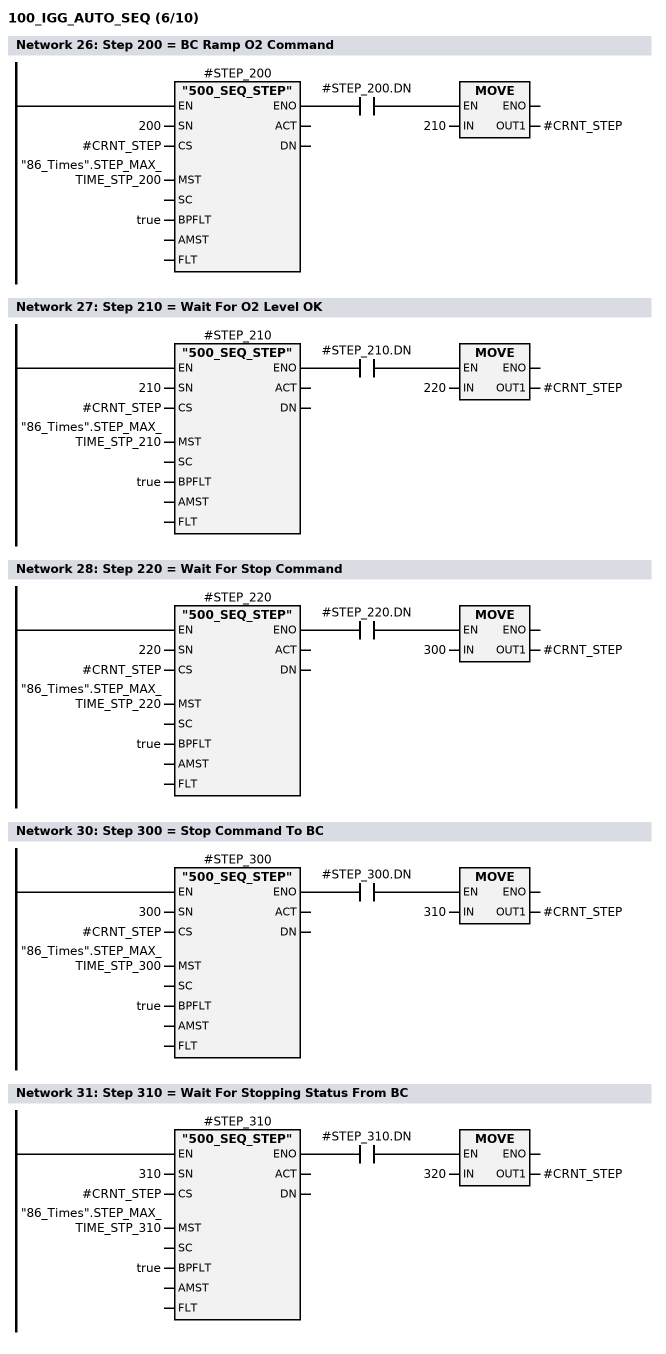
   RUNG wire#powerrail
      #STEP_200(SN := 200, CS := #CRNT_STEP, MST := "86_Times".STEP_MAX_TIME_STP_200, SC :=, BPFLT := true, AMST :=, FLT :=, ACT =>, DN =>)
      Contact( #STEP_200.DN )
      Move(in := 210, out1 => #CRNT_STEP)
   END_RUNG
   // the same network as SCL:
   #STEP_200(SN := 200, CS := #CRNT_STEP, MST := "86_Times".STEP_MAX_TIME_STP_200, BPFLT := true, ENO => #_w1);   // "500_SEQ_STEP"
   IF #_w1 AND #STEP_200.DN THEN #CRNT_STEP := 210; END_IF;
END_REGION

REGION Network 27: Step 210 = Wait For O2 Level OK
   RUNG wire#powerrail
      #STEP_210(SN := 210, CS := #CRNT_STEP, MST := "86_Times".STEP_MAX_TIME_STP_210, SC :=, BPFLT := true, AMST :=, FLT :=, ACT =>, DN =>)
      Contact( #STEP_210.DN )
      Move(in := 220, out1 => #CRNT_STEP)
   END_RUNG
   // the same network as SCL:
   #STEP_210(SN := 210, CS := #CRNT_STEP, MST := "86_Times".STEP_MAX_TIME_STP_210, BPFLT := true, ENO => #_w1);   // "500_SEQ_STEP"
   IF #_w1 AND #STEP_210.DN THEN #CRNT_STEP := 220; END_IF;
END_REGION

REGION Network 28: Step 220 = Wait For Stop Command
   RUNG wire#powerrail
      #STEP_220(SN := 220, CS := #CRNT_STEP, MST := "86_Times".STEP_MAX_TIME_STP_220, SC :=, BPFLT := true, AMST :=, FLT :=, ACT =>, DN =>)
      Contact( #STEP_220.DN )
      Move(in := 300, out1 => #CRNT_STEP)
   END_RUNG
   // the same network as SCL:
   #STEP_220(SN := 220, CS := #CRNT_STEP, MST := "86_Times".STEP_MAX_TIME_STP_220, BPFLT := true, ENO => #_w1);   // "500_SEQ_STEP"
   IF #_w1 AND #STEP_220.DN THEN #CRNT_STEP := 300; END_IF;
END_REGION

REGION Network 30: Step 300 = Stop Command To BC
   RUNG wire#powerrail
      #STEP_300(SN := 300, CS := #CRNT_STEP, MST := "86_Times".STEP_MAX_TIME_STP_300, SC :=, BPFLT := true, AMST :=, FLT :=, ACT =>, DN =>)
      Contact( #STEP_300.DN )
      Move(in := 310, out1 => #CRNT_STEP)
   END_RUNG
   // the same network as SCL:
   #STEP_300(SN := 300, CS := #CRNT_STEP, MST := "86_Times".STEP_MAX_TIME_STP_300, BPFLT := true, ENO => #_w1);   // "500_SEQ_STEP"
   IF #_w1 AND #STEP_300.DN THEN #CRNT_STEP := 310; END_IF;
END_REGION

REGION Network 31: Step 310 = Wait For Stopping Status From BC
   RUNG wire#powerrail
      #STEP_310(SN := 310, CS := #CRNT_STEP, MST := "86_Times".STEP_MAX_TIME_STP_310, SC :=, BPFLT := true, AMST :=, FLT :=, ACT =>, DN =>)
      Contact( #STEP_310.DN )
      Move(in := 320, out1 => #CRNT_STEP)
   END_RUNG
   // the same network as SCL:
   #STEP_310(SN := 310, CS := #CRNT_STEP, MST := "86_Times".STEP_MAX_TIME_STP_310, BPFLT := true, ENO => #_w1);   // "500_SEQ_STEP"
   IF #_w1 AND #STEP_310.DN THEN #CRNT_STEP := 320; END_IF;
END_REGION

REGION Network 32: Step 320 = Wait For O2 Control Stopped From BC
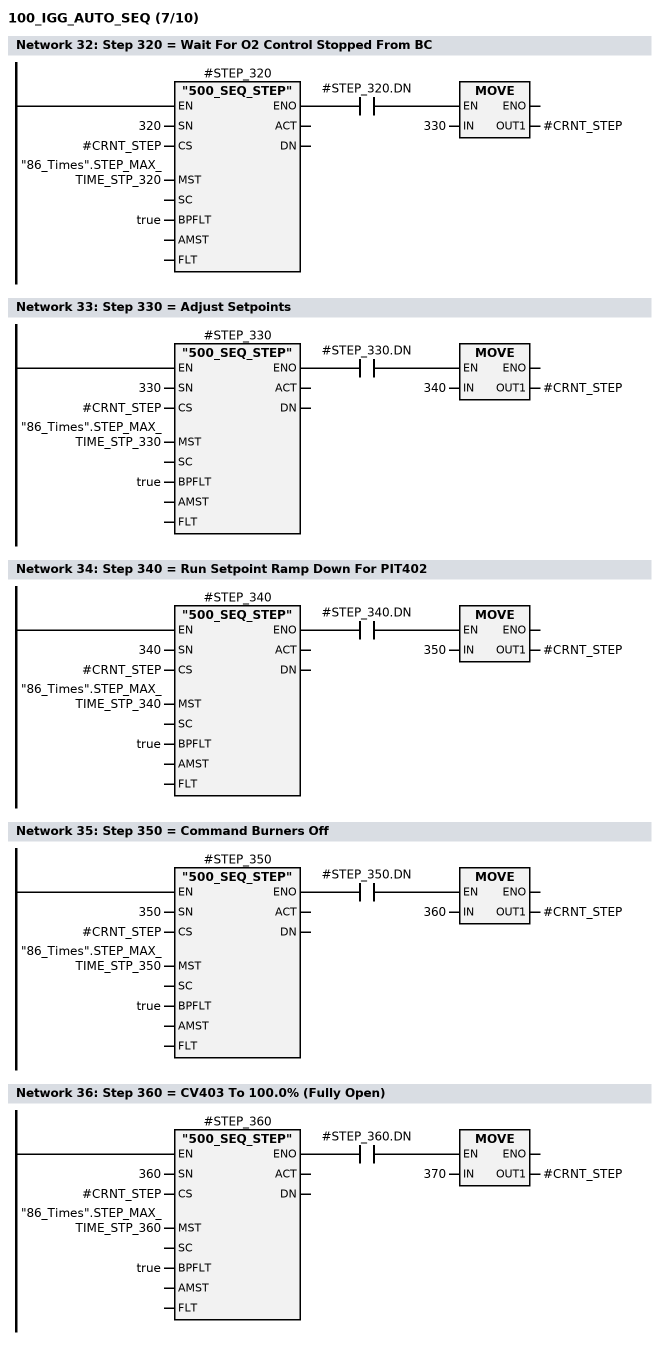
   RUNG wire#powerrail
      #STEP_320(SN := 320, CS := #CRNT_STEP, MST := "86_Times".STEP_MAX_TIME_STP_320, SC :=, BPFLT := true, AMST :=, FLT :=, ACT =>, DN =>)
      Contact( #STEP_320.DN )
      Move(in := 330, out1 => #CRNT_STEP)
   END_RUNG
   // the same network as SCL:
   #STEP_320(SN := 320, CS := #CRNT_STEP, MST := "86_Times".STEP_MAX_TIME_STP_320, BPFLT := true, ENO => #_w1);   // "500_SEQ_STEP"
   IF #_w1 AND #STEP_320.DN THEN #CRNT_STEP := 330; END_IF;
END_REGION

REGION Network 33: Step 330 = Adjust Setpoints
   RUNG wire#powerrail
      #STEP_330(SN := 330, CS := #CRNT_STEP, MST := "86_Times".STEP_MAX_TIME_STP_330, SC :=, BPFLT := true, AMST :=, FLT :=, ACT =>, DN =>)
      Contact( #STEP_330.DN )
      Move(in := 340, out1 => #CRNT_STEP)
   END_RUNG
   // the same network as SCL:
   #STEP_330(SN := 330, CS := #CRNT_STEP, MST := "86_Times".STEP_MAX_TIME_STP_330, BPFLT := true, ENO => #_w1);   // "500_SEQ_STEP"
   IF #_w1 AND #STEP_330.DN THEN #CRNT_STEP := 340; END_IF;
END_REGION

REGION Network 34: Step 340 = Run Setpoint Ramp Down For PIT402
   RUNG wire#powerrail
      #STEP_340(SN := 340, CS := #CRNT_STEP, MST := "86_Times".STEP_MAX_TIME_STP_340, SC :=, BPFLT := true, AMST :=, FLT :=, ACT =>, DN =>)
      Contact( #STEP_340.DN )
      Move(in := 350, out1 => #CRNT_STEP)
   END_RUNG
   // the same network as SCL:
   #STEP_340(SN := 340, CS := #CRNT_STEP, MST := "86_Times".STEP_MAX_TIME_STP_340, BPFLT := true, ENO => #_w1);   // "500_SEQ_STEP"
   IF #_w1 AND #STEP_340.DN THEN #CRNT_STEP := 350; END_IF;
END_REGION

REGION Network 35: Step 350 = Command Burners Off
   RUNG wire#powerrail
      #STEP_350(SN := 350, CS := #CRNT_STEP, MST := "86_Times".STEP_MAX_TIME_STP_350, SC :=, BPFLT := true, AMST :=, FLT :=, ACT =>, DN =>)
      Contact( #STEP_350.DN )
      Move(in := 360, out1 => #CRNT_STEP)
   END_RUNG
   // the same network as SCL:
   #STEP_350(SN := 350, CS := #CRNT_STEP, MST := "86_Times".STEP_MAX_TIME_STP_350, BPFLT := true, ENO => #_w1);   // "500_SEQ_STEP"
   IF #_w1 AND #STEP_350.DN THEN #CRNT_STEP := 360; END_IF;
END_REGION

REGION Network 36: Step 360 = CV403 To 100.0% (Fully Open)
   RUNG wire#powerrail
      #STEP_360(SN := 360, CS := #CRNT_STEP, MST := "86_Times".STEP_MAX_TIME_STP_360, SC :=, BPFLT := true, AMST :=, FLT :=, ACT =>, DN =>)
      Contact( #STEP_360.DN )
      Move(in := 370, out1 => #CRNT_STEP)
   END_RUNG
   // the same network as SCL:
   #STEP_360(SN := 360, CS := #CRNT_STEP, MST := "86_Times".STEP_MAX_TIME_STP_360, BPFLT := true, ENO => #_w1);   // "500_SEQ_STEP"
   IF #_w1 AND #STEP_360.DN THEN #CRNT_STEP := 370; END_IF;
END_REGION

REGION Network 37: Step 370 = Adjust Setpoints
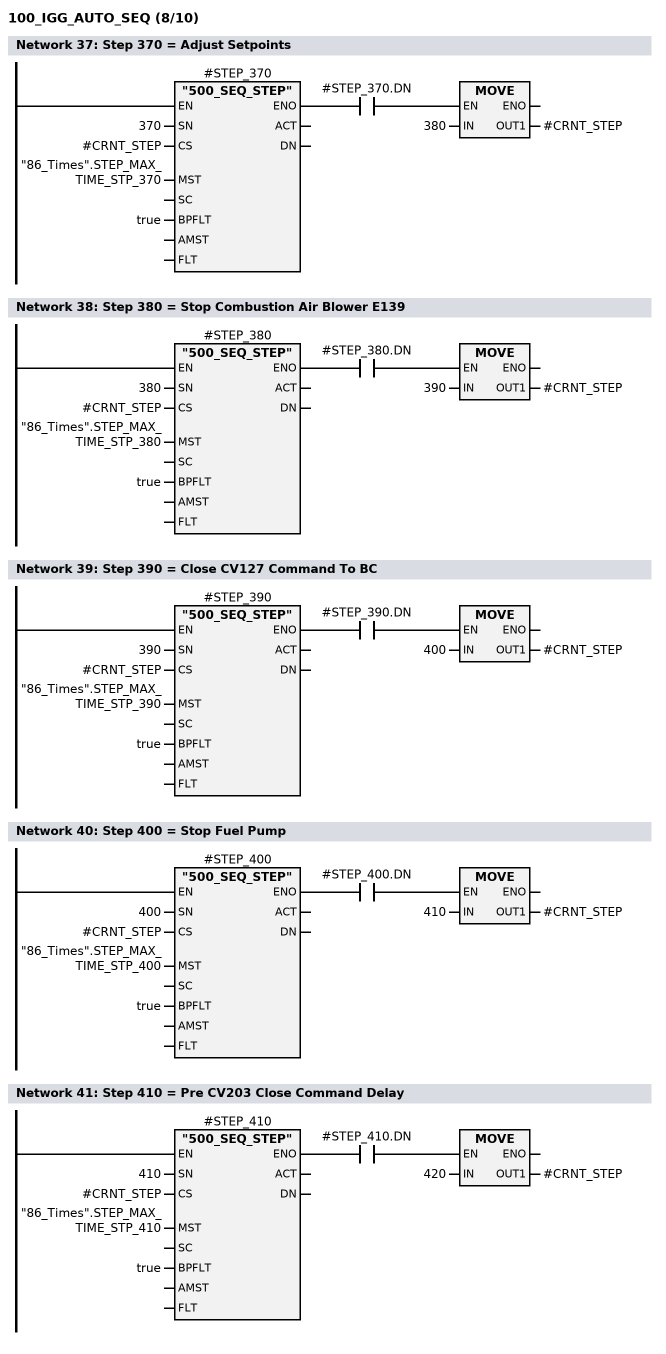
   RUNG wire#powerrail
      #STEP_370(SN := 370, CS := #CRNT_STEP, MST := "86_Times".STEP_MAX_TIME_STP_370, SC :=, BPFLT := true, AMST :=, FLT :=, ACT =>, DN =>)
      Contact( #STEP_370.DN )
      Move(in := 380, out1 => #CRNT_STEP)
   END_RUNG
   // the same network as SCL:
   #STEP_370(SN := 370, CS := #CRNT_STEP, MST := "86_Times".STEP_MAX_TIME_STP_370, BPFLT := true, ENO => #_w1);   // "500_SEQ_STEP"
   IF #_w1 AND #STEP_370.DN THEN #CRNT_STEP := 380; END_IF;
END_REGION

REGION Network 38: Step 380 = Stop Combustion Air Blower E139
   RUNG wire#powerrail
      #STEP_380(SN := 380, CS := #CRNT_STEP, MST := "86_Times".STEP_MAX_TIME_STP_380, SC :=, BPFLT := true, AMST :=, FLT :=, ACT =>, DN =>)
      Contact( #STEP_380.DN )
      Move(in := 390, out1 => #CRNT_STEP)
   END_RUNG
   // the same network as SCL:
   #STEP_380(SN := 380, CS := #CRNT_STEP, MST := "86_Times".STEP_MAX_TIME_STP_380, BPFLT := true, ENO => #_w1);   // "500_SEQ_STEP"
   IF #_w1 AND #STEP_380.DN THEN #CRNT_STEP := 390; END_IF;
END_REGION

REGION Network 39: Step 390 = Close CV127 Command To BC
   RUNG wire#powerrail
      #STEP_390(SN := 390, CS := #CRNT_STEP, MST := "86_Times".STEP_MAX_TIME_STP_390, SC :=, BPFLT := true, AMST :=, FLT :=, ACT =>, DN =>)
      Contact( #STEP_390.DN )
      Move(in := 400, out1 => #CRNT_STEP)
   END_RUNG
   // the same network as SCL:
   #STEP_390(SN := 390, CS := #CRNT_STEP, MST := "86_Times".STEP_MAX_TIME_STP_390, BPFLT := true, ENO => #_w1);   // "500_SEQ_STEP"
   IF #_w1 AND #STEP_390.DN THEN #CRNT_STEP := 400; END_IF;
END_REGION

REGION Network 40: Step 400 = Stop Fuel Pump
   RUNG wire#powerrail
      #STEP_400(SN := 400, CS := #CRNT_STEP, MST := "86_Times".STEP_MAX_TIME_STP_400, SC :=, BPFLT := true, AMST :=, FLT :=, ACT =>, DN =>)
      Contact( #STEP_400.DN )
      Move(in := 410, out1 => #CRNT_STEP)
   END_RUNG
   // the same network as SCL:
   #STEP_400(SN := 400, CS := #CRNT_STEP, MST := "86_Times".STEP_MAX_TIME_STP_400, BPFLT := true, ENO => #_w1);   // "500_SEQ_STEP"
   IF #_w1 AND #STEP_400.DN THEN #CRNT_STEP := 410; END_IF;
END_REGION

REGION Network 41: Step 410 = Pre CV203 Close Command Delay
   RUNG wire#powerrail
      #STEP_410(SN := 410, CS := #CRNT_STEP, MST := "86_Times".STEP_MAX_TIME_STP_410, SC :=, BPFLT := true, AMST :=, FLT :=, ACT =>, DN =>)
      Contact( #STEP_410.DN )
      Move(in := 420, out1 => #CRNT_STEP)
   END_RUNG
   // the same network as SCL:
   #STEP_410(SN := 410, CS := #CRNT_STEP, MST := "86_Times".STEP_MAX_TIME_STP_410, BPFLT := true, ENO => #_w1);   // "500_SEQ_STEP"
   IF #_w1 AND #STEP_410.DN THEN #CRNT_STEP := 420; END_IF;
END_REGION

REGION Network 42: Step 420 = Close CV203 Command To BC
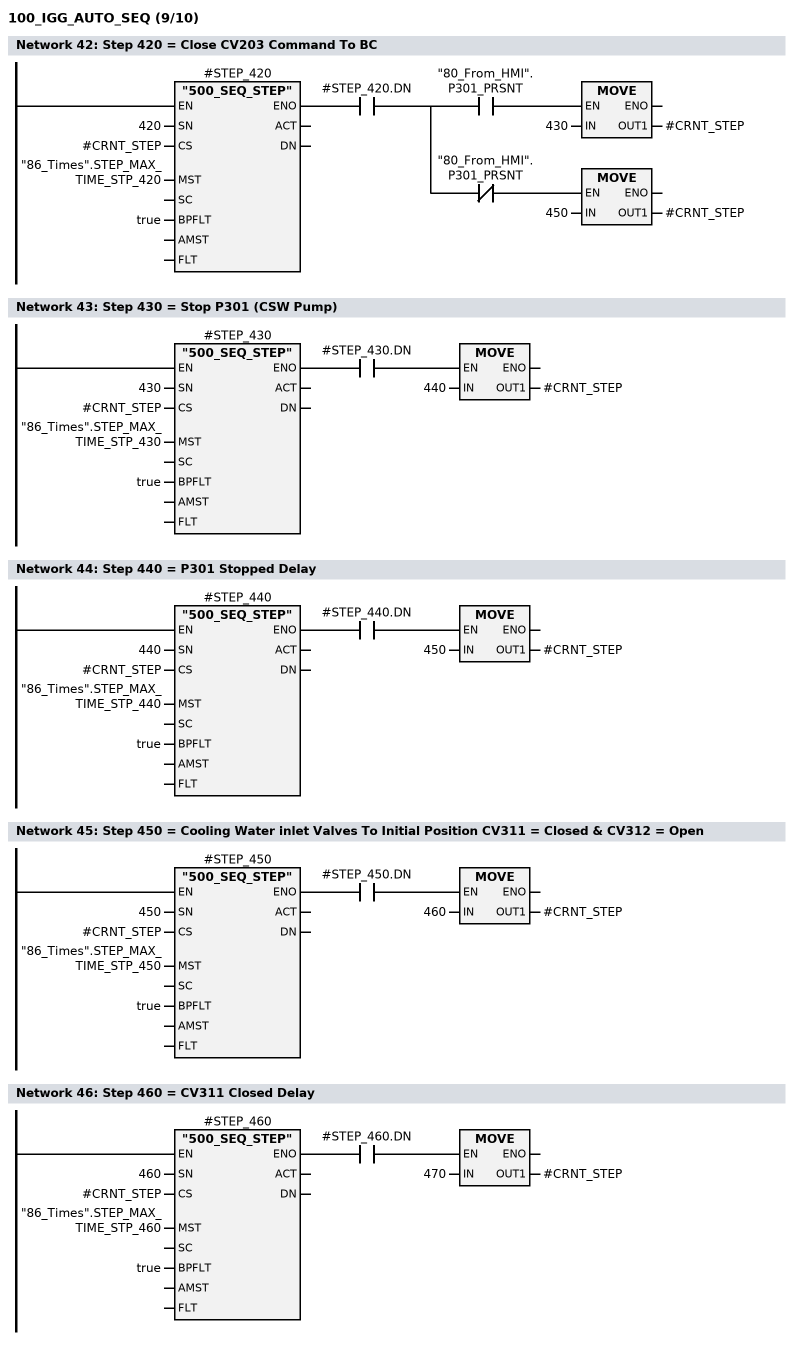
   RUNG wire#powerrail
      #STEP_420(SN := 420, CS := #CRNT_STEP, MST := "86_Times".STEP_MAX_TIME_STP_420, SC :=, BPFLT := true, AMST :=, FLT :=, ACT =>, DN =>)
      Contact( #STEP_420.DN )
      wire#w1
      Contact( "80_From_HMI".P301_PRSNT )
      Move(in := 430, out1 => #CRNT_STEP)
   END_RUNG
   RUNG wire#w1
      I_Contact( "80_From_HMI".P301_PRSNT )
      Move(in := 450, out1 => #CRNT_STEP)
   END_RUNG
   // the same network as SCL:
   #STEP_420(SN := 420, CS := #CRNT_STEP, MST := "86_Times".STEP_MAX_TIME_STP_420, BPFLT := true, ENO => #_w1);   // "500_SEQ_STEP"
   #_w2 := #_w1 AND #STEP_420.DN;
   IF #_w2 AND "80_From_HMI".P301_PRSNT THEN #CRNT_STEP := 430; END_IF;
   IF #_w2 AND NOT "80_From_HMI".P301_PRSNT THEN #CRNT_STEP := 450; END_IF;
END_REGION

REGION Network 43: Step 430 = Stop P301 (CSW Pump)
   RUNG wire#powerrail
      #STEP_430(SN := 430, CS := #CRNT_STEP, MST := "86_Times".STEP_MAX_TIME_STP_430, SC :=, BPFLT := true, AMST :=, FLT :=, ACT =>, DN =>)
      Contact( #STEP_430.DN )
      Move(in := 440, out1 => #CRNT_STEP)
   END_RUNG
   // the same network as SCL:
   #STEP_430(SN := 430, CS := #CRNT_STEP, MST := "86_Times".STEP_MAX_TIME_STP_430, BPFLT := true, ENO => #_w1);   // "500_SEQ_STEP"
   IF #_w1 AND #STEP_430.DN THEN #CRNT_STEP := 440; END_IF;
END_REGION

REGION Network 44: Step 440 = P301 Stopped Delay
   RUNG wire#powerrail
      #STEP_440(SN := 440, CS := #CRNT_STEP, MST := "86_Times".STEP_MAX_TIME_STP_440, SC :=, BPFLT := true, AMST :=, FLT :=, ACT =>, DN =>)
      Contact( #STEP_440.DN )
      Move(in := 450, out1 => #CRNT_STEP)
   END_RUNG
   // the same network as SCL:
   #STEP_440(SN := 440, CS := #CRNT_STEP, MST := "86_Times".STEP_MAX_TIME_STP_440, BPFLT := true, ENO => #_w1);   // "500_SEQ_STEP"
   IF #_w1 AND #STEP_440.DN THEN #CRNT_STEP := 450; END_IF;
END_REGION

REGION Network 45: Step 450 = Cooling Water inlet Valves To Initial Position CV311 = Closed & CV312 = Open
   RUNG wire#powerrail
      #STEP_450(SN := 450, CS := #CRNT_STEP, MST := "86_Times".STEP_MAX_TIME_STP_450, SC :=, BPFLT := true, AMST :=, FLT :=, ACT =>, DN =>)
      Contact( #STEP_450.DN )
      Move(in := 460, out1 => #CRNT_STEP)
   END_RUNG
   // the same network as SCL:
   #STEP_450(SN := 450, CS := #CRNT_STEP, MST := "86_Times".STEP_MAX_TIME_STP_450, BPFLT := true, ENO => #_w1);   // "500_SEQ_STEP"
   IF #_w1 AND #STEP_450.DN THEN #CRNT_STEP := 460; END_IF;
END_REGION

REGION Network 46: Step 460 = CV311 Closed Delay
   RUNG wire#powerrail
      #STEP_460(SN := 460, CS := #CRNT_STEP, MST := "86_Times".STEP_MAX_TIME_STP_460, SC :=, BPFLT := true, AMST :=, FLT :=, ACT =>, DN =>)
      Contact( #STEP_460.DN )
      Move(in := 470, out1 => #CRNT_STEP)
   END_RUNG
   // the same network as SCL:
   #STEP_460(SN := 460, CS := #CRNT_STEP, MST := "86_Times".STEP_MAX_TIME_STP_460, BPFLT := true, ENO => #_w1);   // "500_SEQ_STEP"
   IF #_w1 AND #STEP_460.DN THEN #CRNT_STEP := 470; END_IF;
END_REGION

REGION Network 47: Step 470 = Cooling Water Outlet Valves To Initial Position CV321 = Open & CV322 = Closed
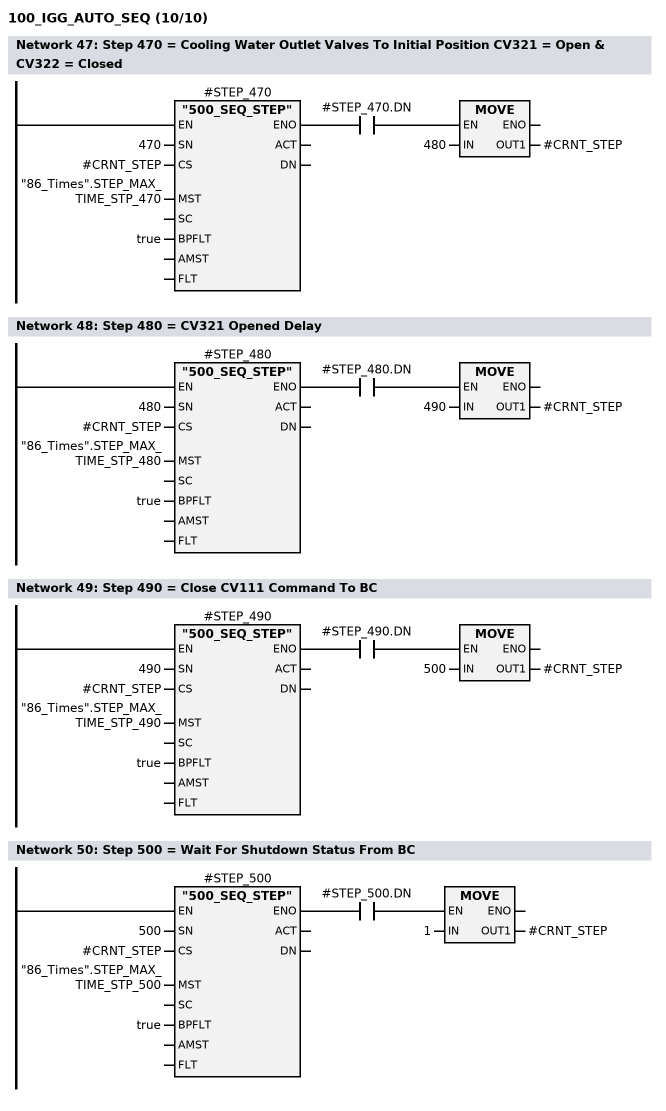
   RUNG wire#powerrail
      #STEP_470(SN := 470, CS := #CRNT_STEP, MST := "86_Times".STEP_MAX_TIME_STP_470, SC :=, BPFLT := true, AMST :=, FLT :=, ACT =>, DN =>)
      Contact( #STEP_470.DN )
      Move(in := 480, out1 => #CRNT_STEP)
   END_RUNG
   // the same network as SCL:
   #STEP_470(SN := 470, CS := #CRNT_STEP, MST := "86_Times".STEP_MAX_TIME_STP_470, BPFLT := true, ENO => #_w1);   // "500_SEQ_STEP"
   IF #_w1 AND #STEP_470.DN THEN #CRNT_STEP := 480; END_IF;
END_REGION

REGION Network 48: Step 480 = CV321 Opened Delay
   RUNG wire#powerrail
      #STEP_480(SN := 480, CS := #CRNT_STEP, MST := "86_Times".STEP_MAX_TIME_STP_480, SC :=, BPFLT := true, AMST :=, FLT :=, ACT =>, DN =>)
      Contact( #STEP_480.DN )
      Move(in := 490, out1 => #CRNT_STEP)
   END_RUNG
   // the same network as SCL:
   #STEP_480(SN := 480, CS := #CRNT_STEP, MST := "86_Times".STEP_MAX_TIME_STP_480, BPFLT := true, ENO => #_w1);   // "500_SEQ_STEP"
   IF #_w1 AND #STEP_480.DN THEN #CRNT_STEP := 490; END_IF;
END_REGION

REGION Network 49: Step 490 = Close CV111 Command To BC
   RUNG wire#powerrail
      #STEP_490(SN := 490, CS := #CRNT_STEP, MST := "86_Times".STEP_MAX_TIME_STP_490, SC :=, BPFLT := true, AMST :=, FLT :=, ACT =>, DN =>)
      Contact( #STEP_490.DN )
      Move(in := 500, out1 => #CRNT_STEP)
   END_RUNG
   // the same network as SCL:
   #STEP_490(SN := 490, CS := #CRNT_STEP, MST := "86_Times".STEP_MAX_TIME_STP_490, BPFLT := true, ENO => #_w1);   // "500_SEQ_STEP"
   IF #_w1 AND #STEP_490.DN THEN #CRNT_STEP := 500; END_IF;
END_REGION

REGION Network 50: Step 500 = Wait For Shutdown Status From BC
   RUNG wire#powerrail
      #STEP_500(SN := 500, CS := #CRNT_STEP, MST := "86_Times".STEP_MAX_TIME_STP_500, SC :=, BPFLT := true, AMST :=, FLT :=, ACT =>, DN =>)
      Contact( #STEP_500.DN )
      Move(in := 1, out1 => #CRNT_STEP)
   END_RUNG
   // the same network as SCL:
   #STEP_500(SN := 500, CS := #CRNT_STEP, MST := "86_Times".STEP_MAX_TIME_STP_500, BPFLT := true, ENO => #_w1);   // "500_SEQ_STEP"
   IF #_w1 AND #STEP_500.DN THEN #CRNT_STEP := 1; END_IF;
END_REGION
END_FUNCTION_BLOCK

FUNCTION_BLOCK "101_Fuel_Pumps"   // FB101, LAD
TITLE = Fuel Pumps Control
{ S7_Optimized_Access := 'TRUE' }
AUTHOR : JRS
VERSION : 0.1
// For the control of duty & standby fuel pumps and associated change over code
   VAR_INPUT
      RUN : Bool;   // Run command
      SW_OVR : Bool;   // Switch pumps request
      "1s_CLK" : Bool;   // 1 Second clock pulse
      MAX_RT : LTime;   // Maximum runtime
      PMP_A_TRP : Bool;   // Pump A tripped
      PMP_A_ENBLD : Bool;   // Pump A running
      PMP_B_TRP : Bool;   // Pump B tripped
      PMP_B_ENBLD : Bool;   // Pump B running
      RST_A_TIM : Bool;   // Reset pump A run time
      RST_B_TIM : Bool;   // Reset pump B run time
   END_VAR
   VAR_OUTPUT
      RUN_A : Bool;   // Run pump A
      RUN_B : Bool;   // Run pump B
   END_VAR
   VAR_IN_OUT
      "Run Time A" : LTime;   // Pump A current run time
      "Run Time B" : LTime;   // Pump B current run time
      "Duty Is A" : Bool;   // Duty bit
      "Duty Is B" : Bool;   // Duty bit
   END_VAR
   VAR
      "A Pulse Bit" : Bool;   // Pulse bit
      "B Pulse Bit" : Bool;   // Pulse bit
      "SW Pulse Bit" : Bool;   // Pulse bit
      "SW Pulse Bit_N" : Bool;
      "SW Latch" : Bool;   // Switch over latch bit
      "SW Latch_Manual" : Bool;
      Aux1 : Bool;
   END_VAR
   VAR_TEMP   // added for the SCL form of the ladder/FBD networks
      _w1 : Bool;
      _w2 : Bool;
      _w3 : Bool;
   END_VAR
BEGIN

REGION Network 1: Pump A Run Time
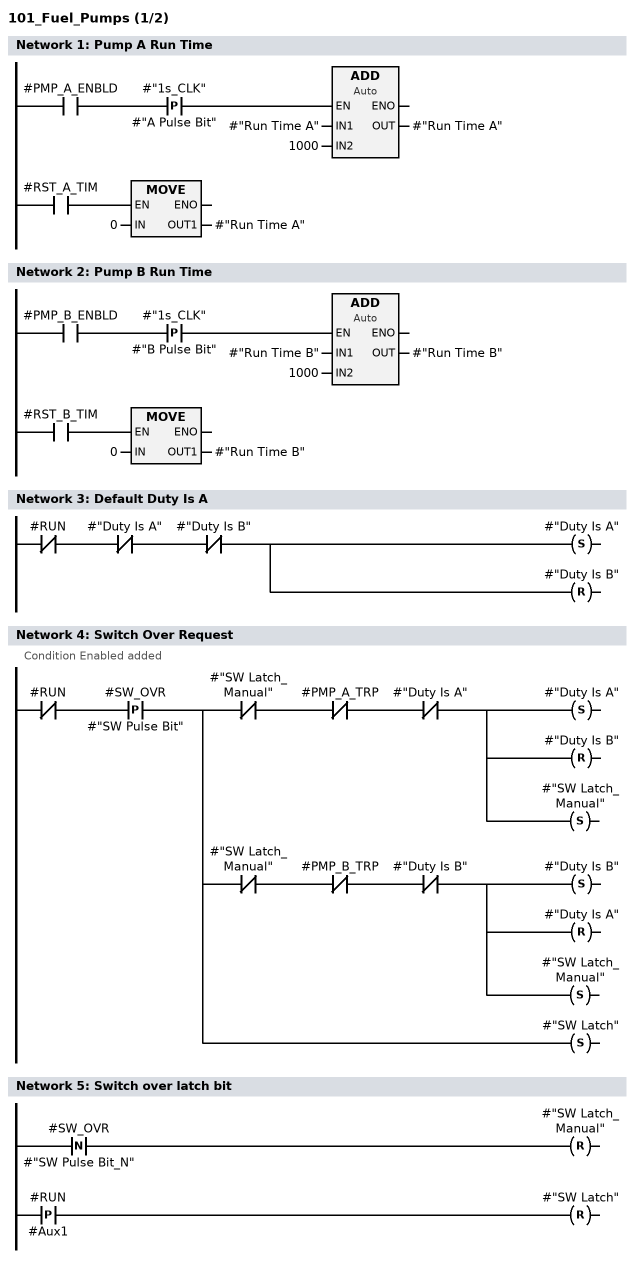
   RUNG wire#powerrail
      Contact( #PMP_A_ENBLD )
      P_Contact(operand := #"1s_CLK", bit := #"A Pulse Bit")
      Add(in1 := #"Run Time A", in2 := 1000, out => #"Run Time A")
   END_RUNG
   RUNG wire#powerrail
      Contact( #RST_A_TIM )
      Move(in := 0, out1 => #"Run Time A")
   END_RUNG
   // the same network as SCL:
   #_w1 := #PMP_A_ENBLD AND #"1s_CLK" AND NOT #"A Pulse Bit";   // rising edge of #"1s_CLK"
   #"A Pulse Bit" := #"1s_CLK";
   IF #_w1 THEN #"Run Time A" := #"Run Time A" + 1000; END_IF;
   IF #RST_A_TIM THEN #"Run Time A" := 0; END_IF;
END_REGION

REGION Network 2: Pump B Run Time
   RUNG wire#powerrail
      Contact( #PMP_B_ENBLD )
      P_Contact(operand := #"1s_CLK", bit := #"B Pulse Bit")
      Add(in1 := #"Run Time B", in2 := 1000, out => #"Run Time B")
   END_RUNG
   RUNG wire#powerrail
      Contact( #RST_B_TIM )
      Move(in := 0, out1 => #"Run Time B")
   END_RUNG
   // the same network as SCL:
   #_w1 := #PMP_B_ENBLD AND #"1s_CLK" AND NOT #"B Pulse Bit";   // rising edge of #"1s_CLK"
   #"B Pulse Bit" := #"1s_CLK";
   IF #_w1 THEN #"Run Time B" := #"Run Time B" + 1000; END_IF;
   IF #RST_B_TIM THEN #"Run Time B" := 0; END_IF;
END_REGION

REGION Network 3: Default Duty Is A
   RUNG wire#powerrail
      I_Contact( #RUN )
      I_Contact( #"Duty Is A" )
      I_Contact( #"Duty Is B" )
      wire#w1
      S_Coil( #"Duty Is A" )
   END_RUNG
   RUNG wire#w1
      R_Coil( #"Duty Is B" )
   END_RUNG
   // the same network as SCL:
   #_w1 := NOT #RUN AND NOT #"Duty Is A" AND NOT #"Duty Is B";
   IF #_w1 THEN
       #"Duty Is A" := TRUE;
       #"Duty Is B" := FALSE;
   END_IF;
END_REGION

REGION Network 4: Switch Over Request
   // Condition Enabled added
   RUNG wire#powerrail
      I_Contact( #RUN )
      P_Contact(operand := #SW_OVR, bit := #"SW Pulse Bit")
      wire#w1
      I_Contact( #"SW Latch_Manual" )
      I_Contact( #PMP_A_TRP )
      I_Contact( #"Duty Is A" )
      wire#w2
      S_Coil( #"Duty Is A" )
   END_RUNG
   RUNG wire#w2
      R_Coil( #"Duty Is B" )
   END_RUNG
   RUNG wire#w2
      S_Coil( #"SW Latch_Manual" )
   END_RUNG
   RUNG wire#w1
      I_Contact( #"SW Latch_Manual" )
      I_Contact( #PMP_B_TRP )
      I_Contact( #"Duty Is B" )
      wire#w3
      S_Coil( #"Duty Is B" )
   END_RUNG
   RUNG wire#w3
      R_Coil( #"Duty Is A" )
   END_RUNG
   RUNG wire#w3
      S_Coil( #"SW Latch_Manual" )
   END_RUNG
   RUNG wire#w1
      S_Coil( #"SW Latch" )
   END_RUNG
   // the same network as SCL:
   #_w1 := NOT #RUN AND #SW_OVR AND NOT #"SW Pulse Bit";   // rising edge of #SW_OVR
   #"SW Pulse Bit" := #SW_OVR;
   #_w2 := #_w1 AND NOT #"SW Latch_Manual" AND NOT #PMP_A_TRP AND NOT #"Duty Is A";
   IF #_w2 THEN
       #"Duty Is A" := TRUE;
       #"Duty Is B" := FALSE;
       #"SW Latch_Manual" := TRUE;
   END_IF;
   #_w3 := #_w1 AND NOT #"SW Latch_Manual" AND NOT #PMP_B_TRP AND NOT #"Duty Is B";
   IF #_w3 THEN
       #"Duty Is B" := TRUE;
       #"Duty Is A" := FALSE;
       #"SW Latch_Manual" := TRUE;
   END_IF;
   IF #_w1 THEN #"SW Latch" := TRUE; END_IF;
END_REGION

REGION Network 5: Switch over latch bit
   RUNG wire#powerrail
      N_Contact(operand := #SW_OVR, bit := #"SW Pulse Bit_N")
      R_Coil( #"SW Latch_Manual" )
   END_RUNG
   RUNG wire#powerrail
      P_Contact(operand := #RUN, bit := #Aux1)
      R_Coil( #"SW Latch" )
   END_RUNG
   // the same network as SCL:
   #_w1 := NOT #SW_OVR AND #"SW Pulse Bit_N";   // falling edge of #SW_OVR
   #"SW Pulse Bit_N" := #SW_OVR;
   IF #_w1 THEN #"SW Latch_Manual" := FALSE; END_IF;
   #_w2 := #RUN AND NOT #Aux1;   // rising edge of #RUN
   #Aux1 := #RUN;
   IF #_w2 THEN #"SW Latch" := FALSE; END_IF;
END_REGION

REGION Network 6: Auto Change To A
   // Changed to change to A on B tripped during work.
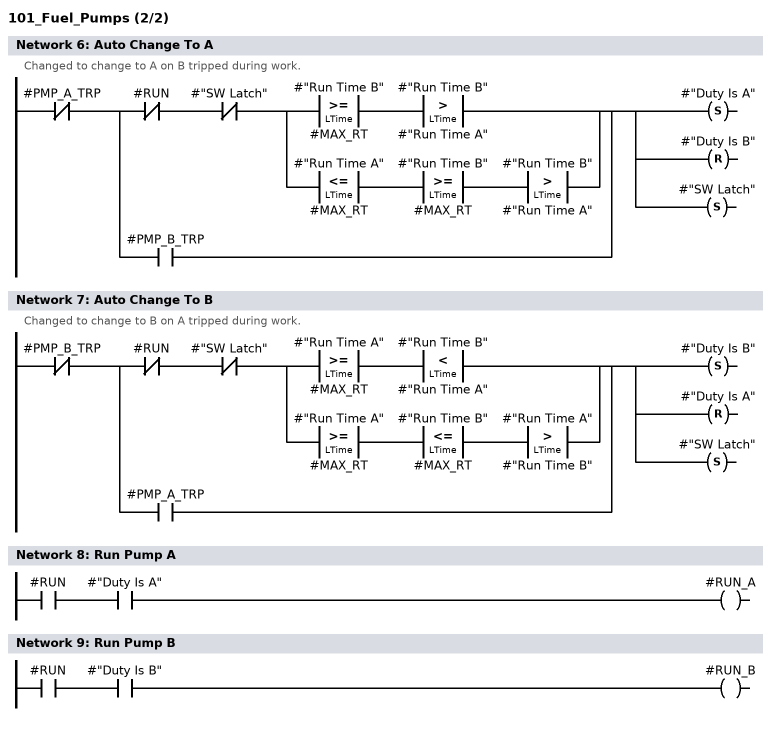
   RUNG wire#powerrail
      I_Contact( #PMP_A_TRP )
      wire#w1
      I_Contact( #RUN )
      I_Contact( #"SW Latch" )
      wire#w2
      { S7_Templates := "SrcType := LTime" } GE_Contact(in1 := #"Run Time B", in2 := #MAX_RT)
      { S7_Templates := "SrcType := LTime" } GT_Contact(in1 := #"Run Time B", in2 := #"Run Time A")
      wire#w3
      S_Coil( #"Duty Is A" )
   END_RUNG
   RUNG wire#w2
      { S7_Templates := "SrcType := LTime" } LE_Contact(in1 := #"Run Time A", in2 := #MAX_RT)
      { S7_Templates := "SrcType := LTime" } GE_Contact(in1 := #"Run Time B", in2 := #MAX_RT)
      { S7_Templates := "SrcType := LTime" } GT_Contact(in1 := #"Run Time B", in2 := #"Run Time A")
   END_RUNG wire#w3
   RUNG wire#w1
      Contact( #PMP_B_TRP )
   END_RUNG wire#w3
   RUNG wire#w3
      R_Coil( #"Duty Is B" )
   END_RUNG
   RUNG wire#w3
      S_Coil( #"SW Latch" )
   END_RUNG
   // the same network as SCL:
   IF NOT #PMP_A_TRP AND ((NOT #RUN AND NOT #"SW Latch" AND (((#"Run Time B" >= #MAX_RT) AND (#"Run Time B" > #"Run Time A")) OR ((#"Run Time A" <= #MAX_RT) AND (#"Run Time B" >= #MAX_RT) AND (#"Run Time B" > #"Run Time A")))) OR #PMP_B_TRP) THEN
       #"Duty Is A" := TRUE;
       #"Duty Is B" := FALSE;
       #"SW Latch" := TRUE;
   END_IF;
END_REGION

REGION Network 7: Auto Change To B
   // Changed to change to B on A tripped during work.
   RUNG wire#powerrail
      I_Contact( #PMP_B_TRP )
      wire#w1
      I_Contact( #RUN )
      I_Contact( #"SW Latch" )
      wire#w2
      { S7_Templates := "SrcType := LTime" } GE_Contact(in1 := #"Run Time A", in2 := #MAX_RT)
      { S7_Templates := "SrcType := LTime" } LT_Contact(in1 := #"Run Time B", in2 := #"Run Time A")
      wire#w3
      S_Coil( #"Duty Is B" )
   END_RUNG
   RUNG wire#w2
      { S7_Templates := "SrcType := LTime" } GE_Contact(in1 := #"Run Time A", in2 := #MAX_RT)
      { S7_Templates := "SrcType := LTime" } LE_Contact(in1 := #"Run Time B", in2 := #MAX_RT)
      { S7_Templates := "SrcType := LTime" } GT_Contact(in1 := #"Run Time A", in2 := #"Run Time B")
   END_RUNG wire#w3
   RUNG wire#w1
      Contact( #PMP_A_TRP )
   END_RUNG wire#w3
   RUNG wire#w3
      R_Coil( #"Duty Is A" )
   END_RUNG
   RUNG wire#w3
      S_Coil( #"SW Latch" )
   END_RUNG
   // the same network as SCL:
   IF NOT #PMP_B_TRP AND ((NOT #RUN AND NOT #"SW Latch" AND (((#"Run Time A" >= #MAX_RT) AND (#"Run Time B" < #"Run Time A")) OR ((#"Run Time A" >= #MAX_RT) AND (#"Run Time B" <= #MAX_RT) AND (#"Run Time A" > #"Run Time B")))) OR #PMP_A_TRP) THEN
       #"Duty Is B" := TRUE;
       #"Duty Is A" := FALSE;
       #"SW Latch" := TRUE;
   END_IF;
END_REGION

REGION Network 8: Run Pump A
   RUNG wire#powerrail
      Contact( #RUN )
      Contact( #"Duty Is A" )
      Coil( #RUN_A )
   END_RUNG
   // the same network as SCL:
   #RUN_A := #RUN AND #"Duty Is A";
END_REGION

REGION Network 9: Run Pump B
   RUNG wire#powerrail
      Contact( #RUN )
      Contact( #"Duty Is B" )
      Coil( #RUN_B )
   END_RUNG
   // the same network as SCL:
   #RUN_B := #RUN AND #"Duty Is B";
END_REGION
END_FUNCTION_BLOCK

FUNCTION_BLOCK "105_SP_RAMP_PIT402_UP"   // FB105, LAD
TITLE = Setpoint Ramp Up For PIT402
{ S7_Optimized_Access := 'TRUE' }
AUTHOR : JRS
VERSION : 0.1
// Determines the live setpoint value for PIT402 based on target and ramp time
   VAR_INPUT
      RUN : Bool;   // Demand
      INIT_SP : Real;   // Initial setpoint
      TRGT_SP : Real;   // Target setpoint
      RMP_SECS : Int := 30;   // To target ramp time in seconds
      "1Hz_PULSE" : Bool;   // 1 Hz clock pulse
      RST : Bool;   // Reset flag
   END_VAR
   VAR_OUTPUT
      DN : Bool;   // Done
      FLT : Bool;   // Fault
   END_VAR
   VAR_IN_OUT
      RUNNING : Bool;   // Block is running
      TARGET : Real;   // Target
   END_VAR
   VAR
      STATE : Int;   // State value
      INTO_RUN_EDGE : Bool;   // Edge bit
      OUT_OF_RUN_EDGE : Bool;   // Edge bit
      RST_FLG : Bool;   // Reset flag
      PS_STP_VAL : Real;   // Per second step value
      CLK_PLS_EDGE : Bool;   // Clock pulse edge
      IEC_Timer_0_Instance : TON_TIME;
   END_VAR
   VAR_TEMP   // added for the SCL form of the ladder/FBD networks
      _w1 : Bool;
   END_VAR
BEGIN

REGION Network 1: Running
   // For running status detection
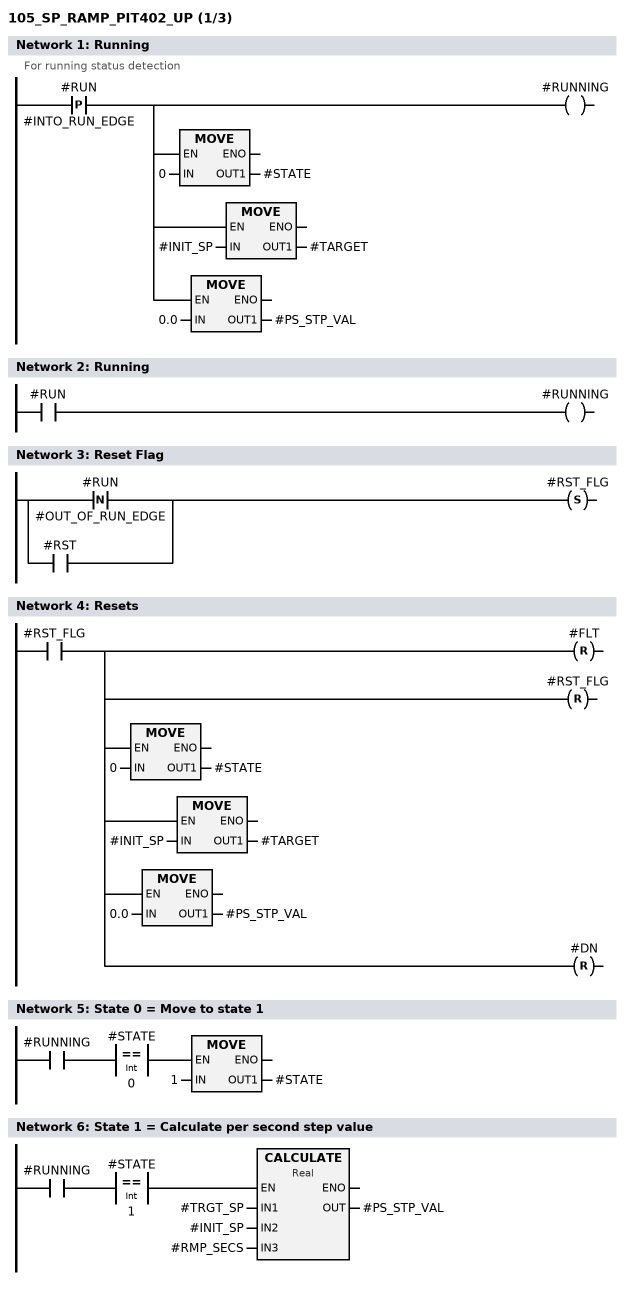
   RUNG wire#powerrail
      P_Contact(operand := #RUN, bit := #INTO_RUN_EDGE)
      wire#w1
      Coil( #RUNNING )
   END_RUNG
   RUNG wire#w1
      Move(in := 0, out1 => #STATE)
   END_RUNG
   RUNG wire#w1
      Move(in := #INIT_SP, out1 => #TARGET)
   END_RUNG
   RUNG wire#w1
      Move(in := 0.0, out1 => #PS_STP_VAL)
   END_RUNG
   // the same network as SCL:
   #_w1 := #RUN AND NOT #INTO_RUN_EDGE;   // rising edge of #RUN
   #INTO_RUN_EDGE := #RUN;
   #RUNNING := #_w1;
   IF #_w1 THEN
       #STATE := 0;
       #TARGET := #INIT_SP;
       #PS_STP_VAL := 0.0;
   END_IF;
END_REGION

REGION Network 2: Running
   RUNG wire#powerrail
      Contact( #RUN )
      Coil( #RUNNING )
   END_RUNG
   // the same network as SCL:
   #RUNNING := #RUN;
END_REGION

REGION Network 3: Reset Flag
   RUNG wire#powerrail
      N_Contact(operand := #RUN, bit := #OUT_OF_RUN_EDGE)
      wire#w1
      S_Coil( #RST_FLG )
   END_RUNG
   RUNG wire#powerrail
      Contact( #RST )
   END_RUNG wire#w1
   // the same network as SCL:
   #_w1 := NOT #RUN AND #OUT_OF_RUN_EDGE;   // falling edge of #RUN
   #OUT_OF_RUN_EDGE := #RUN;
   IF #_w1 OR #RST THEN #RST_FLG := TRUE; END_IF;
END_REGION

REGION Network 4: Resets
   RUNG wire#powerrail
      Contact( #RST_FLG )
      wire#w1
      R_Coil( #FLT )
   END_RUNG
   RUNG wire#w1
      R_Coil( #RST_FLG )
   END_RUNG
   RUNG wire#w1
      Move(in := 0, out1 => #STATE)
   END_RUNG
   RUNG wire#w1
      Move(in := #INIT_SP, out1 => #TARGET)
   END_RUNG
   RUNG wire#w1
      Move(in := 0.0, out1 => #PS_STP_VAL)
   END_RUNG
   RUNG wire#w1
      R_Coil( #DN )
   END_RUNG
   // the same network as SCL:
   IF #RST_FLG THEN #FLT := FALSE; END_IF;
   #_w1 := #RST_FLG;
   IF #_w1 THEN
       #RST_FLG := FALSE;
       #STATE := 0;
       #TARGET := #INIT_SP;
       #PS_STP_VAL := 0.0;
       #DN := FALSE;
   END_IF;
END_REGION

REGION Network 5: State 0 = Move to state 1
   RUNG wire#powerrail
      Contact( #RUNNING )
      { S7_Templates := "SrcType := Int" } EQ_Contact(in1 := #STATE, in2 := 0)
      Move(in := 1, out1 => #STATE)
   END_RUNG
   // the same network as SCL:
   IF #RUNNING AND (#STATE = 0) THEN #STATE := 1; END_IF;
END_REGION

REGION Network 6: State 1 = Calculate per second step value
   RUNG wire#powerrail
      Contact( #RUNNING )
      { S7_Templates := "SrcType := Int" } EQ_Contact(in1 := #STATE, in2 := 1)
      { S7_Templates := "SrcType := Real"; S7_Expression := "(IN1-IN2)/IN3" } Calculate(in1 := #TRGT_SP, in2 := #INIT_SP, in3 := #RMP_SECS, out => #PS_STP_VAL)
   END_RUNG
   // the same network as SCL:
   IF #RUNNING AND (#STATE = 1) THEN #PS_STP_VAL := (#TRGT_SP-#INIT_SP)/#RMP_SECS; END_IF;
END_REGION

REGION Network 7: Into State 2
